   RUNG wire#w1
      R_Coil( %DB60.DBX2.7 )
   END_RUNG
   RUNG wire#w1
      R_Coil( %DB60.DBX3.0 )
   END_RUNG
   RUNG wire#w1
      R_Coil( %DB60.DBX3.1 )
   END_RUNG
   RUNG wire#w1
      R_Coil( %DB60.DBX3.2 )
   END_RUNG
   RUNG wire#w1
      R_Coil( %DB60.DBX3.3 )
   END_RUNG
   RUNG wire#w1
      R_Coil( %DB60.DBX3.4 )
   END_RUNG
   RUNG wire#w1
      R_Coil( %DB60.DBX3.5 )
   END_RUNG
   RUNG wire#w1
      R_Coil( %DB60.DBX3.6 )
   END_RUNG
   RUNG wire#w1
      R_Coil( %DB60.DBX3.7 )
   END_RUNG
   RUNG wire#w1
      R_Coil( %DB60.DBX4.0 )
   END_RUNG
   RUNG wire#w1
      R_Coil( %DB60.DBX4.1 )
   END_RUNG
   RUNG wire#w1
      R_Coil( %DB60.DBX4.2 )
   END_RUNG
   RUNG wire#w1
      R_Coil( %DB60.DBX4.3 )
   END_RUNG
   RUNG wire#w1
      R_Coil( %DB60.DBX4.4 )
   END_RUNG
   RUNG wire#w1
      R_Coil( %DB60.DBX4.5 )
   END_RUNG
   RUNG wire#w1
      R_Coil( %DB60.DBX4.6 )
   END_RUNG
   RUNG wire#w1
      R_Coil( %DB60.DBX4.7 )
   END_RUNG
   RUNG wire#w1
      R_Coil( %DB60.DBX5.0 )
   END_RUNG
   RUNG wire#w1
      R_Coil( %DB60.DBX5.1 )
   END_RUNG
   RUNG wire#w1
      R_Coil( %DB60.DBX5.2 )
   END_RUNG
   RUNG wire#w1
      R_Coil( %DB60.DBX5.3 )
   END_RUNG
   RUNG wire#w1
      R_Coil( %DB60.DBX5.4 )
   END_RUNG
   RUNG wire#w1
      R_Coil( %DB60.DBX5.5 )
   END_RUNG
   RUNG wire#w1
      R_Coil( %DB60.DBX5.6 )
   END_RUNG
   RUNG wire#w1
      R_Coil( %DB60.DBX5.7 )
   END_RUNG
   RUNG wire#w1
      R_Coil( %DB60.DBX6.0 )
   END_RUNG
   RUNG wire#w1
      R_Coil( %DB60.DBX6.1 )
   END_RUNG
   RUNG wire#w1
      R_Coil( %DB60.DBX6.2 )
   END_RUNG
   RUNG wire#w1
      R_Coil( %DB60.DBX6.3 )
   END_RUNG
   RUNG wire#w1
      R_Coil( %DB60.DBX6.4 )
   END_RUNG
   RUNG wire#w1
      R_Coil( %DB60.DBX6.5 )
   END_RUNG
   RUNG wire#w1
      R_Coil( %DB60.DBX6.6 )
   END_RUNG
   RUNG wire#w1
      R_Coil( %DB60.DBX6.7 )
   END_RUNG
   RUNG wire#w1
      R_Coil( %DB60.DBX7.0 )
   END_RUNG
   RUNG wire#w1
      R_Coil( %DB60.DBX7.1 )
   END_RUNG
   RUNG wire#w1
      R_Coil( %DB60.DBX7.2 )
   END_RUNG
   RUNG wire#w1
      R_Coil( %DB60.DBX7.3 )
   END_RUNG
   RUNG wire#w1
      R_Coil( %DB60.DBX7.4 )
   END_RUNG
   RUNG wire#w1
      R_Coil( %DB60.DBX7.5 )
   END_RUNG
   RUNG wire#w1
      R_Coil( %DB60.DBX7.6 )
   END_RUNG
   RUNG wire#w1
      R_Coil( %DB60.DBX7.7 )
   END_RUNG
   // the same network as SCL:
   IF "50_CMND_DATA".Alarm_Reset THEN
       %DB60.DBX0.0 := FALSE;
       %DB60.DBX0.1 := FALSE;
       %DB60.DBX0.2 := FALSE;
       %DB60.DBX0.3 := FALSE;
       %DB60.DBX0.4 := FALSE;
       %DB60.DBX0.5 := FALSE;
       %DB60.DBX0.6 := FALSE;
       %DB60.DBX0.7 := FALSE;
       %DB60.DBX1.0 := FALSE;
       %DB60.DBX1.1 := FALSE;
       %DB60.DBX1.2 := FALSE;
       %DB60.DBX1.3 := FALSE;
       %DB60.DBX1.4 := FALSE;
       %DB60.DBX1.5 := FALSE;
       %DB60.DBX1.6 := FALSE;
       %DB60.DBX1.7 := FALSE;
       %DB60.DBX2.0 := FALSE;
       %DB60.DBX2.1 := FALSE;
       %DB60.DBX2.2 := FALSE;
       %DB60.DBX2.3 := FALSE;
       %DB60.DBX2.4 := FALSE;
       %DB60.DBX2.5 := FALSE;
       %DB60.DBX2.6 := FALSE;
       %DB60.DBX2.7 := FALSE;
       %DB60.DBX3.0 := FALSE;
       %DB60.DBX3.1 := FALSE;
       %DB60.DBX3.2 := FALSE;
       %DB60.DBX3.3 := FALSE;
       %DB60.DBX3.4 := FALSE;
       %DB60.DBX3.5 := FALSE;
       %DB60.DBX3.6 := FALSE;
       %DB60.DBX3.7 := FALSE;
       %DB60.DBX4.0 := FALSE;
       %DB60.DBX4.1 := FALSE;
       %DB60.DBX4.2 := FALSE;
       %DB60.DBX4.3 := FALSE;
       %DB60.DBX4.4 := FALSE;
       %DB60.DBX4.5 := FALSE;
       %DB60.DBX4.6 := FALSE;
       %DB60.DBX4.7 := FALSE;
       %DB60.DBX5.0 := FALSE;
       %DB60.DBX5.1 := FALSE;
       %DB60.DBX5.2 := FALSE;
       %DB60.DBX5.3 := FALSE;
       %DB60.DBX5.4 := FALSE;
       %DB60.DBX5.5 := FALSE;
       %DB60.DBX5.6 := FALSE;
       %DB60.DBX5.7 := FALSE;
       %DB60.DBX6.0 := FALSE;
       %DB60.DBX6.1 := FALSE;
       %DB60.DBX6.2 := FALSE;
       %DB60.DBX6.3 := FALSE;
       %DB60.DBX6.4 := FALSE;
       %DB60.DBX6.5 := FALSE;
       %DB60.DBX6.6 := FALSE;
       %DB60.DBX6.7 := FALSE;
       %DB60.DBX7.0 := FALSE;
       %DB60.DBX7.1 := FALSE;
       %DB60.DBX7.2 := FALSE;
       %DB60.DBX7.3 := FALSE;
       %DB60.DBX7.4 := FALSE;
       %DB60.DBX7.5 := FALSE;
       %DB60.DBX7.6 := FALSE;
       %DB60.DBX7.7 := FALSE;
   END_IF;
END_REGION

REGION Network 34: Alarm Present
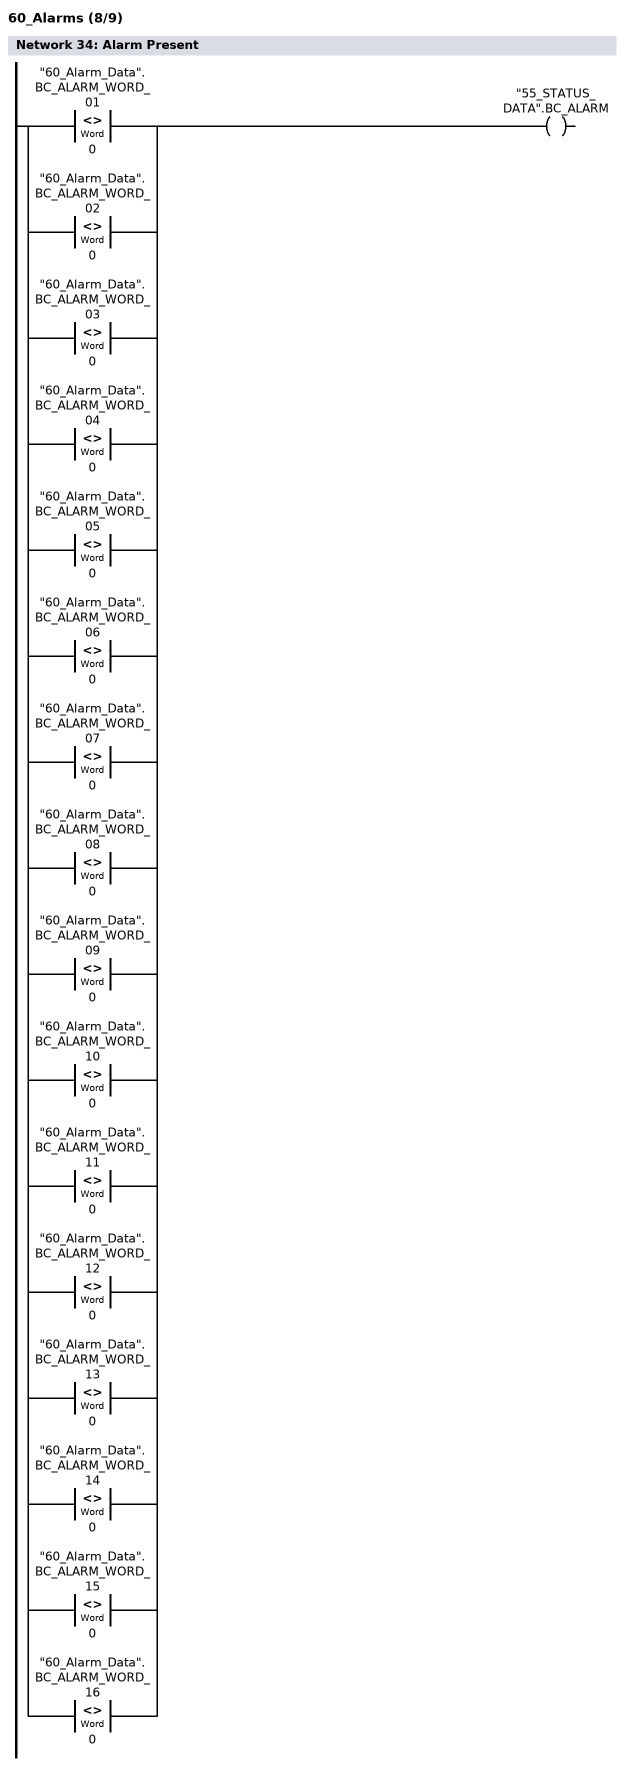
   RUNG wire#powerrail
      { S7_Templates := "SrcType := Word" } NE_Contact(in1 := "60_Alarm_Data".BC_ALARM_WORD_01, in2 := 0)
      wire#w1
      Coil( "55_STATUS_DATA".BC_ALARM )
   END_RUNG
   RUNG wire#powerrail
      { S7_Templates := "SrcType := Word" } NE_Contact(in1 := "60_Alarm_Data".BC_ALARM_WORD_02, in2 := 0)
   END_RUNG wire#w1
   RUNG wire#powerrail
      { S7_Templates := "SrcType := Word" } NE_Contact(in1 := "60_Alarm_Data".BC_ALARM_WORD_03, in2 := 0)
   END_RUNG wire#w1
   RUNG wire#powerrail
      { S7_Templates := "SrcType := Word" } NE_Contact(in1 := "60_Alarm_Data".BC_ALARM_WORD_04, in2 := 0)
   END_RUNG wire#w1
   RUNG wire#powerrail
      { S7_Templates := "SrcType := Word" } NE_Contact(in1 := "60_Alarm_Data".BC_ALARM_WORD_05, in2 := 0)
   END_RUNG wire#w1
   RUNG wire#powerrail
      { S7_Templates := "SrcType := Word" } NE_Contact(in1 := "60_Alarm_Data".BC_ALARM_WORD_06, in2 := 0)
   END_RUNG wire#w1
   RUNG wire#powerrail
      { S7_Templates := "SrcType := Word" } NE_Contact(in1 := "60_Alarm_Data".BC_ALARM_WORD_07, in2 := 0)
   END_RUNG wire#w1
   RUNG wire#powerrail
      { S7_Templates := "SrcType := Word" } NE_Contact(in1 := "60_Alarm_Data".BC_ALARM_WORD_08, in2 := 0)
   END_RUNG wire#w1
   RUNG wire#powerrail
      { S7_Templates := "SrcType := Word" } NE_Contact(in1 := "60_Alarm_Data".BC_ALARM_WORD_09, in2 := 0)
   END_RUNG wire#w1
   RUNG wire#powerrail
      { S7_Templates := "SrcType := Word" } NE_Contact(in1 := "60_Alarm_Data".BC_ALARM_WORD_10, in2 := 0)
   END_RUNG wire#w1
   RUNG wire#powerrail
      { S7_Templates := "SrcType := Word" } NE_Contact(in1 := "60_Alarm_Data".BC_ALARM_WORD_11, in2 := 0)
   END_RUNG wire#w1
   RUNG wire#powerrail
      { S7_Templates := "SrcType := Word" } NE_Contact(in1 := "60_Alarm_Data".BC_ALARM_WORD_12, in2 := 0)
   END_RUNG wire#w1
   RUNG wire#powerrail
      { S7_Templates := "SrcType := Word" } NE_Contact(in1 := "60_Alarm_Data".BC_ALARM_WORD_13, in2 := 0)
   END_RUNG wire#w1
   RUNG wire#powerrail
      { S7_Templates := "SrcType := Word" } NE_Contact(in1 := "60_Alarm_Data".BC_ALARM_WORD_14, in2 := 0)
   END_RUNG wire#w1
   RUNG wire#powerrail
      { S7_Templates := "SrcType := Word" } NE_Contact(in1 := "60_Alarm_Data".BC_ALARM_WORD_15, in2 := 0)
   END_RUNG wire#w1
   RUNG wire#powerrail
      { S7_Templates := "SrcType := Word" } NE_Contact(in1 := "60_Alarm_Data".BC_ALARM_WORD_16, in2 := 0)
   END_RUNG wire#w1
   // the same network as SCL:
   "55_STATUS_DATA".BC_ALARM := ("60_Alarm_Data".BC_ALARM_WORD_01 <> 0) OR ("60_Alarm_Data".BC_ALARM_WORD_02 <> 0) OR ("60_Alarm_Data".BC_ALARM_WORD_03 <> 0) OR ("60_Alarm_Data".BC_ALARM_WORD_04 <> 0) OR ("60_Alarm_Data".BC_ALARM_WORD_05 <> 0) OR ("60_Alarm_Data".BC_ALARM_WORD_06 <> 0) OR ("60_Alarm_Data".BC_ALARM_WORD_07 <> 0) OR ("60_Alarm_Data".BC_ALARM_WORD_08 <> 0) OR ("60_Alarm_Data".BC_ALARM_WORD_09 <> 0) OR ("60_Alarm_Data".BC_ALARM_WORD_10 <> 0) OR ("60_Alarm_Data".BC_ALARM_WORD_11 <> 0) OR ("60_Alarm_Data".BC_ALARM_WORD_12 <> 0) OR ("60_Alarm_Data".BC_ALARM_WORD_13 <> 0) OR ("60_Alarm_Data".BC_ALARM_WORD_14 <> 0) OR ("60_Alarm_Data".BC_ALARM_WORD_15 <> 0) OR ("60_Alarm_Data".BC_ALARM_WORD_16 <> 0);
END_REGION

REGION Network 35: Alarm present
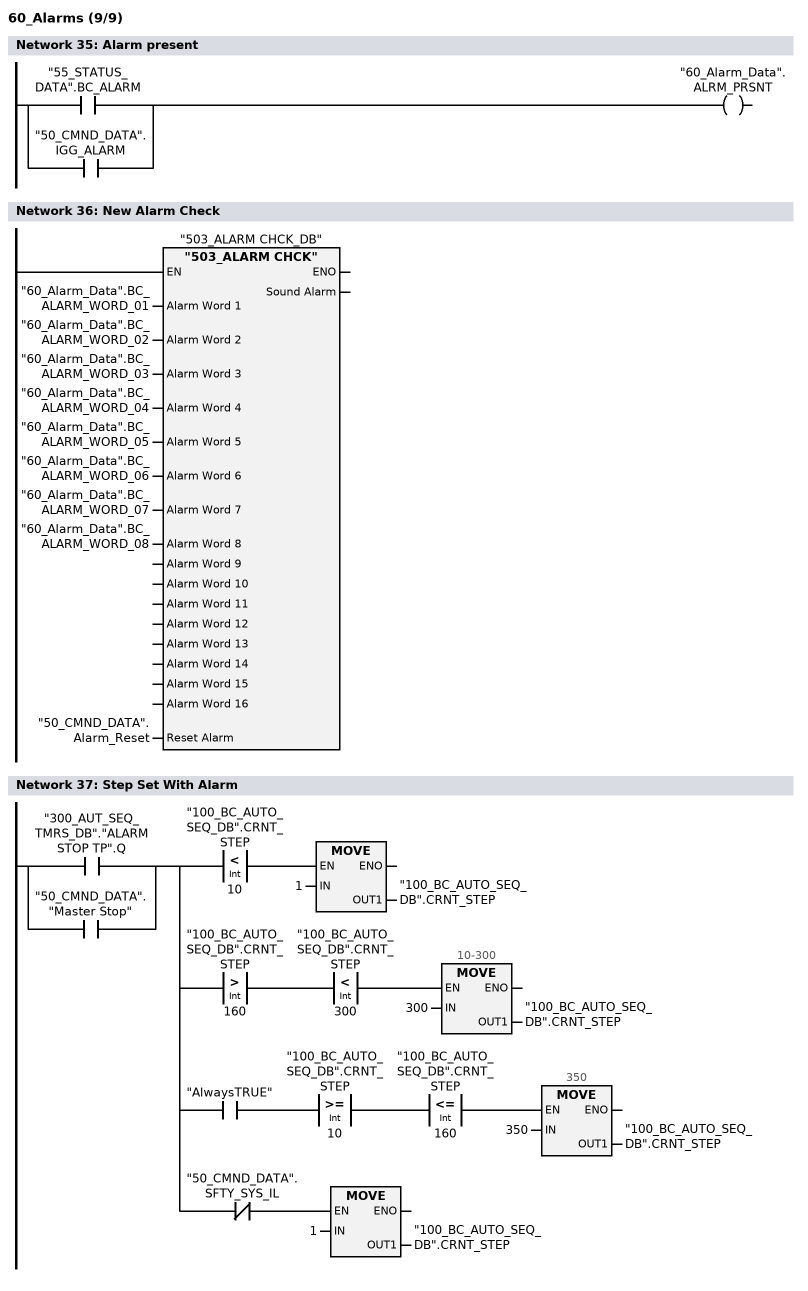
   RUNG wire#powerrail
      Contact( "55_STATUS_DATA".BC_ALARM )
      wire#w1
      Coil( "60_Alarm_Data".ALRM_PRSNT )
   END_RUNG
   RUNG wire#powerrail
      Contact( "50_CMND_DATA".IGG_ALARM )
   END_RUNG wire#w1
   // the same network as SCL:
   "60_Alarm_Data".ALRM_PRSNT := "55_STATUS_DATA".BC_ALARM OR "50_CMND_DATA".IGG_ALARM;
END_REGION

REGION Network 36: New Alarm Check
   RUNG wire#powerrail
      "503_ALARM CHCK_DB"("Alarm Word 1" := "60_Alarm_Data".BC_ALARM_WORD_01, "Alarm Word 2" := "60_Alarm_Data".BC_ALARM_WORD_02, "Alarm Word 3" := "60_Alarm_Data".BC_ALARM_WORD_03, "Alarm Word 4" := "60_Alarm_Data".BC_ALARM_WORD_04, "Alarm Word 5" := "60_Alarm_Data".BC_ALARM_WORD_05, "Alarm Word 6" := "60_Alarm_Data".BC_ALARM_WORD_06, "Alarm Word 7" := "60_Alarm_Data".BC_ALARM_WORD_07, "Alarm Word 8" := "60_Alarm_Data".BC_ALARM_WORD_08, "Alarm Word 9" :=, "Alarm Word 10" :=, "Alarm Word 11" :=, "Alarm Word 12" :=, "Alarm Word 13" :=, "Alarm Word 14" :=, "Alarm Word 15" :=, "Alarm Word 16" :=, "Reset Alarm" := "50_CMND_DATA".Alarm_Reset, "Sound Alarm" =>)
   END_RUNG
   // the same network as SCL:
   "503_ALARM CHCK_DB"("Alarm Word 1" := "60_Alarm_Data".BC_ALARM_WORD_01,   // "503_ALARM CHCK"
                       "Alarm Word 2" := "60_Alarm_Data".BC_ALARM_WORD_02,
                       "Alarm Word 3" := "60_Alarm_Data".BC_ALARM_WORD_03,
                       "Alarm Word 4" := "60_Alarm_Data".BC_ALARM_WORD_04,
                       "Alarm Word 5" := "60_Alarm_Data".BC_ALARM_WORD_05,
                       "Alarm Word 6" := "60_Alarm_Data".BC_ALARM_WORD_06,
                       "Alarm Word 7" := "60_Alarm_Data".BC_ALARM_WORD_07,
                       "Alarm Word 8" := "60_Alarm_Data".BC_ALARM_WORD_08,
                       "Reset Alarm" := "50_CMND_DATA".Alarm_Reset);
END_REGION

REGION Network 37: Step Set With Alarm
   RUNG wire#powerrail
      Contact( "300_AUT_SEQ_TMRS_DB"."ALARM STOP TP".Q )
      wire#w1
      { S7_Templates := "SrcType := Int" } LT_Contact(in1 := "100_BC_AUTO_SEQ_DB".CRNT_STEP, in2 := 10)
      Move(in := 1, out1 => "100_BC_AUTO_SEQ_DB".CRNT_STEP)
   END_RUNG
   RUNG wire#powerrail
      Contact( "50_CMND_DATA"."Master Stop" )
   END_RUNG wire#w1
   RUNG wire#w1
      { S7_Templates := "SrcType := Int" } GT_Contact(in1 := "100_BC_AUTO_SEQ_DB".CRNT_STEP, in2 := 160)
      { S7_Templates := "SrcType := Int" } LT_Contact(in1 := "100_BC_AUTO_SEQ_DB".CRNT_STEP, in2 := 300)
      Move(in := 300, out1 => "100_BC_AUTO_SEQ_DB".CRNT_STEP)   // 10-300
   END_RUNG
   RUNG wire#w1
      Contact( "AlwaysTRUE" )
      { S7_Templates := "SrcType := Int" } GE_Contact(in1 := "100_BC_AUTO_SEQ_DB".CRNT_STEP, in2 := 10)
      { S7_Templates := "SrcType := Int" } LE_Contact(in1 := "100_BC_AUTO_SEQ_DB".CRNT_STEP, in2 := 160)
      Move(in := 350, out1 => "100_BC_AUTO_SEQ_DB".CRNT_STEP)   // 350
   END_RUNG
   RUNG wire#w1
      I_Contact( "50_CMND_DATA".SFTY_SYS_IL )
      Move(in := 1, out1 => "100_BC_AUTO_SEQ_DB".CRNT_STEP)
   END_RUNG
   // the same network as SCL:
   #_w1 := "300_AUT_SEQ_TMRS_DB"."ALARM STOP TP".Q OR "50_CMND_DATA"."Master Stop";
   IF #_w1 AND ("100_BC_AUTO_SEQ_DB".CRNT_STEP < 10) THEN "100_BC_AUTO_SEQ_DB".CRNT_STEP := 1; END_IF;
   IF #_w1 AND ("100_BC_AUTO_SEQ_DB".CRNT_STEP > 160) AND ("100_BC_AUTO_SEQ_DB".CRNT_STEP < 300) THEN
       "100_BC_AUTO_SEQ_DB".CRNT_STEP := 300;   // 10-300
   END_IF;
   IF #_w1 AND "AlwaysTRUE" AND ("100_BC_AUTO_SEQ_DB".CRNT_STEP >= 10) AND ("100_BC_AUTO_SEQ_DB".CRNT_STEP <= 160) THEN
       "100_BC_AUTO_SEQ_DB".CRNT_STEP := 350;   // 350
   END_IF;
   IF #_w1 AND NOT "50_CMND_DATA".SFTY_SYS_IL THEN "100_BC_AUTO_SEQ_DB".CRNT_STEP := 1; END_IF;
END_REGION
END_FUNCTION

FUNCTION "62_Warnings" : Void   // FC62, LAD
TITLE = Warning Processing
{ S7_Optimized_Access := 'TRUE' }
AUTHOR : JRS
VERSION : 0.1
// To warning conditions
   VAR_TEMP   // added for the SCL form of the ladder/FBD networks
      _w1 : Bool;
   END_VAR
BEGIN

REGION Network 1: DB62 WORD_1 =PIT204 Fuel Oil pessure transmitter
   // BC_WARNING_WORD_01 BIT 1/2/3/4
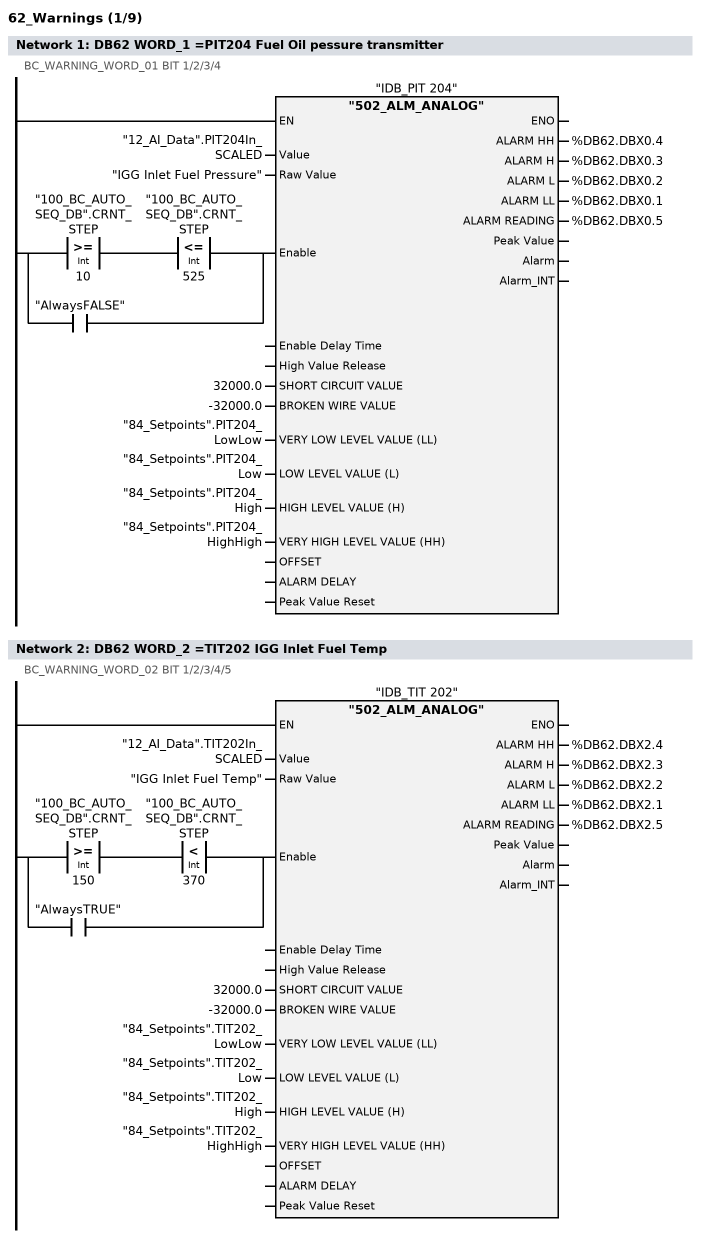
   RUNG wire#powerrail
      "IDB_PIT 204"(Enable := wire#w1, Value := "12_AI_Data".PIT204In_SCALED, "Raw Value" := "IGG Inlet Fuel Pressure", "SHORT CIRCUIT VALUE" := 32000.0, "BROKEN WIRE VALUE" := -32000.0, "VERY LOW LEVEL VALUE (LL)" := "84_Setpoints".PIT204_LowLow, "LOW LEVEL VALUE (L)" := "84_Setpoints".PIT204_Low, "HIGH LEVEL VALUE (H)" := "84_Setpoints".PIT204_High, "VERY HIGH LEVEL VALUE (HH)" := "84_Setpoints".PIT204_HighHigh, OFFSET :=, "ALARM DELAY" :=, "Peak Value Reset" :=, "ALARM HH" => %DB62.DBX0.4, "ALARM H" => %DB62.DBX0.3, "ALARM L" => %DB62.DBX0.2, "ALARM LL" => %DB62.DBX0.1, "ALARM READING" => %DB62.DBX0.5, "Peak Value" =>, Alarm =>, Alarm_INT =>, "Enable Delay Time" :=, "High Value Release" :=)
   END_RUNG
   RUNG wire#powerrail
      { S7_Templates := "SrcType := Int" } GE_Contact(in1 := "100_BC_AUTO_SEQ_DB".CRNT_STEP, in2 := 10)
      { S7_Templates := "SrcType := Int" } LE_Contact(in1 := "100_BC_AUTO_SEQ_DB".CRNT_STEP, in2 := 525)
   END_RUNG wire#w1
   RUNG wire#powerrail
      Contact( "AlwaysFALSE" )
   END_RUNG wire#w1
   // the same network as SCL:
   "IDB_PIT 204"(Value := "12_AI_Data".PIT204In_SCALED,   // "502_ALM_ANALOG"
                 "Raw Value" := "IGG Inlet Fuel Pressure",
                 Enable := (("100_BC_AUTO_SEQ_DB".CRNT_STEP >= 10) AND ("100_BC_AUTO_SEQ_DB".CRNT_STEP <= 525)) OR "AlwaysFALSE",
                 "SHORT CIRCUIT VALUE" := 32000.0,
                 "BROKEN WIRE VALUE" := -32000.0,
                 "VERY LOW LEVEL VALUE (LL)" := "84_Setpoints".PIT204_LowLow,
                 "LOW LEVEL VALUE (L)" := "84_Setpoints".PIT204_Low,
                 "HIGH LEVEL VALUE (H)" := "84_Setpoints".PIT204_High,
                 "VERY HIGH LEVEL VALUE (HH)" := "84_Setpoints".PIT204_HighHigh,
                 "ALARM HH" => %DB62.DBX0.4,
                 "ALARM H" => %DB62.DBX0.3,
                 "ALARM L" => %DB62.DBX0.2,
                 "ALARM LL" => %DB62.DBX0.1,
                 "ALARM READING" => %DB62.DBX0.5);
END_REGION

REGION Network 2: DB62 WORD_2 =TIT202 IGG Inlet Fuel Temp
   // BC_WARNING_WORD_02 BIT 1/2/3/4/5
   RUNG wire#powerrail
      "IDB_TIT 202"(Enable := wire#w1, Value := "12_AI_Data".TIT202In_SCALED, "Raw Value" := "IGG Inlet Fuel Temp", "SHORT CIRCUIT VALUE" := 32000.0, "BROKEN WIRE VALUE" := -32000.0, "VERY LOW LEVEL VALUE (LL)" := "84_Setpoints".TIT202_LowLow, "LOW LEVEL VALUE (L)" := "84_Setpoints".TIT202_Low, "HIGH LEVEL VALUE (H)" := "84_Setpoints".TIT202_High, "VERY HIGH LEVEL VALUE (HH)" := "84_Setpoints".TIT202_HighHigh, OFFSET :=, "ALARM DELAY" :=, "Peak Value Reset" :=, "ALARM HH" => %DB62.DBX2.4, "ALARM H" => %DB62.DBX2.3, "ALARM L" => %DB62.DBX2.2, "ALARM LL" => %DB62.DBX2.1, "ALARM READING" => %DB62.DBX2.5, "Peak Value" =>, Alarm =>, Alarm_INT =>, "Enable Delay Time" :=, "High Value Release" :=)
   END_RUNG
   RUNG wire#powerrail
      { S7_Templates := "SrcType := Int" } GE_Contact(in1 := "100_BC_AUTO_SEQ_DB".CRNT_STEP, in2 := 150)
      { S7_Templates := "SrcType := Int" } LT_Contact(in1 := "100_BC_AUTO_SEQ_DB".CRNT_STEP, in2 := 370)
   END_RUNG wire#w1
   RUNG wire#powerrail
      Contact( "AlwaysTRUE" )
   END_RUNG wire#w1
   // the same network as SCL:
   "IDB_TIT 202"(Value := "12_AI_Data".TIT202In_SCALED,   // "502_ALM_ANALOG"
                 "Raw Value" := "IGG Inlet Fuel Temp",
                 Enable := (("100_BC_AUTO_SEQ_DB".CRNT_STEP >= 150) AND ("100_BC_AUTO_SEQ_DB".CRNT_STEP < 370)) OR "AlwaysTRUE",
                 "SHORT CIRCUIT VALUE" := 32000.0,
                 "BROKEN WIRE VALUE" := -32000.0,
                 "VERY LOW LEVEL VALUE (LL)" := "84_Setpoints".TIT202_LowLow,
                 "LOW LEVEL VALUE (L)" := "84_Setpoints".TIT202_Low,
                 "HIGH LEVEL VALUE (H)" := "84_Setpoints".TIT202_High,
                 "VERY HIGH LEVEL VALUE (HH)" := "84_Setpoints".TIT202_HighHigh,
                 "ALARM HH" => %DB62.DBX2.4,
                 "ALARM H" => %DB62.DBX2.3,
                 "ALARM L" => %DB62.DBX2.2,
                 "ALARM LL" => %DB62.DBX2.1,
                 "ALARM READING" => %DB62.DBX2.5);
END_REGION

REGION Network 3: DB62 WORD_3 =PIT205 IGG Main Fuel Pressure
   // BC_WARNING_WORD_03
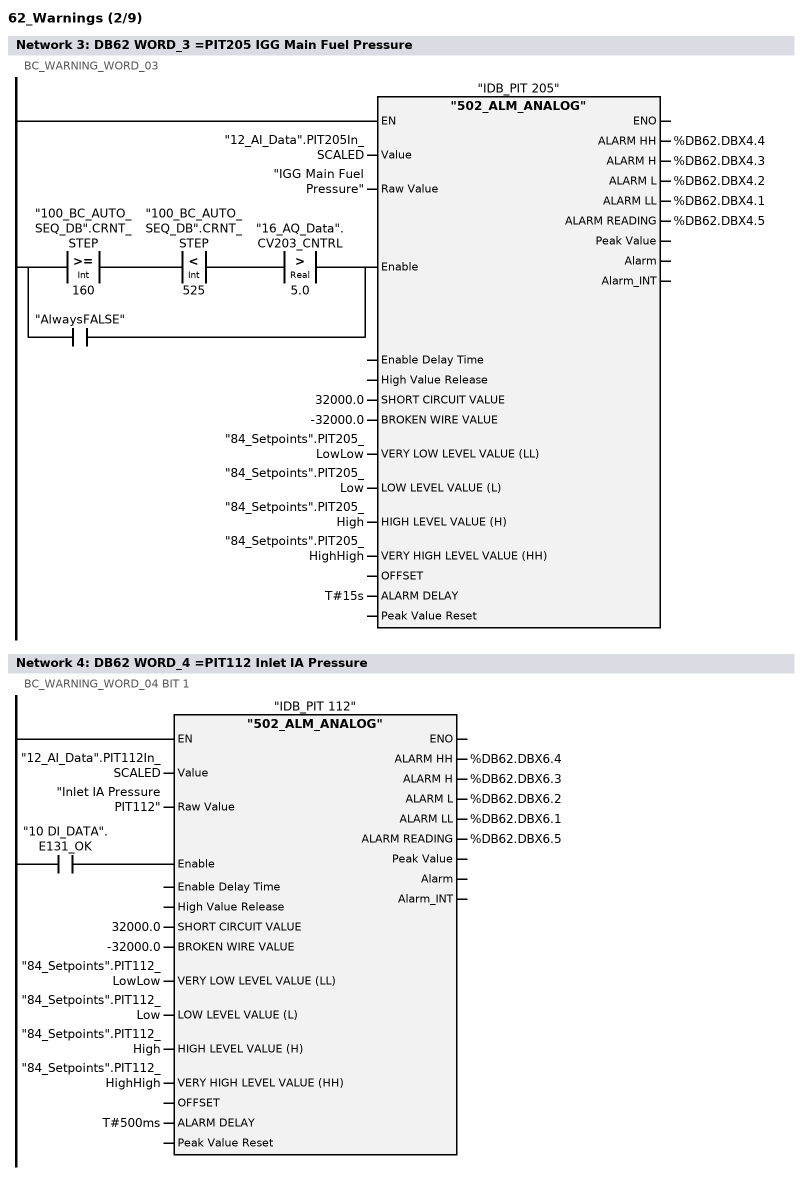
   RUNG wire#powerrail
      "IDB_PIT 205"(Enable := wire#w1, Value := "12_AI_Data".PIT205In_SCALED, "Raw Value" := "IGG Main Fuel Pressure", "SHORT CIRCUIT VALUE" := 32000.0, "BROKEN WIRE VALUE" := -32000.0, "VERY LOW LEVEL VALUE (LL)" := "84_Setpoints".PIT205_LowLow, "LOW LEVEL VALUE (L)" := "84_Setpoints".PIT205_Low, "HIGH LEVEL VALUE (H)" := "84_Setpoints".PIT205_High, "VERY HIGH LEVEL VALUE (HH)" := "84_Setpoints".PIT205_HighHigh, OFFSET :=, "ALARM DELAY" := T#15s, "Peak Value Reset" :=, "ALARM HH" => %DB62.DBX4.4, "ALARM H" => %DB62.DBX4.3, "ALARM L" => %DB62.DBX4.2, "ALARM LL" => %DB62.DBX4.1, "ALARM READING" => %DB62.DBX4.5, "Peak Value" =>, Alarm =>, Alarm_INT =>, "Enable Delay Time" :=, "High Value Release" :=)
   END_RUNG
   RUNG wire#powerrail
      { S7_Templates := "SrcType := Int" } GE_Contact(in1 := "100_BC_AUTO_SEQ_DB".CRNT_STEP, in2 := 160)
      { S7_Templates := "SrcType := Int" } LT_Contact(in1 := "100_BC_AUTO_SEQ_DB".CRNT_STEP, in2 := 525)
      { S7_Templates := "SrcType := Real" } GT_Contact(in1 := "16_AQ_Data".CV203_CNTRL, in2 := 5.0)
   END_RUNG wire#w1
   RUNG wire#powerrail
      Contact( "AlwaysFALSE" )
   END_RUNG wire#w1
   // the same network as SCL:
   "IDB_PIT 205"(Value := "12_AI_Data".PIT205In_SCALED,   // "502_ALM_ANALOG"
                 "Raw Value" := "IGG Main Fuel Pressure",
                 Enable := (("100_BC_AUTO_SEQ_DB".CRNT_STEP >= 160) AND ("100_BC_AUTO_SEQ_DB".CRNT_STEP < 525) AND ("16_AQ_Data".CV203_CNTRL > 5.0)) OR "AlwaysFALSE",
                 "SHORT CIRCUIT VALUE" := 32000.0,
                 "BROKEN WIRE VALUE" := -32000.0,
                 "VERY LOW LEVEL VALUE (LL)" := "84_Setpoints".PIT205_LowLow,
                 "LOW LEVEL VALUE (L)" := "84_Setpoints".PIT205_Low,
                 "HIGH LEVEL VALUE (H)" := "84_Setpoints".PIT205_High,
                 "VERY HIGH LEVEL VALUE (HH)" := "84_Setpoints".PIT205_HighHigh,
                 "ALARM DELAY" := T#15s,
                 "ALARM HH" => %DB62.DBX4.4,
                 "ALARM H" => %DB62.DBX4.3,
                 "ALARM L" => %DB62.DBX4.2,
                 "ALARM LL" => %DB62.DBX4.1,
                 "ALARM READING" => %DB62.DBX4.5);
END_REGION

REGION Network 4: DB62 WORD_4 =PIT112 Inlet IA Pressure
   // BC_WARNING_WORD_04 BIT 1
   RUNG wire#powerrail
      "IDB_PIT 112"(Enable := wire#w1, Value := "12_AI_Data".PIT112In_SCALED, "Raw Value" := "Inlet IA Pressure PIT112", "SHORT CIRCUIT VALUE" := 32000.0, "BROKEN WIRE VALUE" := -32000.0, "VERY LOW LEVEL VALUE (LL)" := "84_Setpoints".PIT112_LowLow, "LOW LEVEL VALUE (L)" := "84_Setpoints".PIT112_Low, "HIGH LEVEL VALUE (H)" := "84_Setpoints".PIT112_High, "VERY HIGH LEVEL VALUE (HH)" := "84_Setpoints".PIT112_HighHigh, OFFSET :=, "ALARM DELAY" := T#500ms, "Peak Value Reset" :=, "ALARM HH" => %DB62.DBX6.4, "ALARM H" => %DB62.DBX6.3, "ALARM L" => %DB62.DBX6.2, "ALARM LL" => %DB62.DBX6.1, "ALARM READING" => %DB62.DBX6.5, "Peak Value" =>, Alarm =>, Alarm_INT =>, "Enable Delay Time" :=, "High Value Release" :=)
   END_RUNG
   RUNG wire#powerrail
      Contact( "10 DI_DATA".E131_OK )
   END_RUNG wire#w1
   // the same network as SCL:
   "IDB_PIT 112"(Value := "12_AI_Data".PIT112In_SCALED,   // "502_ALM_ANALOG"
                 "Raw Value" := "Inlet IA Pressure PIT112",
                 Enable := "10 DI_DATA".E131_OK,
                 "SHORT CIRCUIT VALUE" := 32000.0,
                 "BROKEN WIRE VALUE" := -32000.0,
                 "VERY LOW LEVEL VALUE (LL)" := "84_Setpoints".PIT112_LowLow,
                 "LOW LEVEL VALUE (L)" := "84_Setpoints".PIT112_Low,
                 "HIGH LEVEL VALUE (H)" := "84_Setpoints".PIT112_High,
                 "VERY HIGH LEVEL VALUE (HH)" := "84_Setpoints".PIT112_HighHigh,
                 "ALARM DELAY" := T#500ms,
                 "ALARM HH" => %DB62.DBX6.4,
                 "ALARM H" => %DB62.DBX6.3,
                 "ALARM L" => %DB62.DBX6.2,
                 "ALARM LL" => %DB62.DBX6.1,
                 "ALARM READING" => %DB62.DBX6.5);
END_REGION

REGION Network 5: DB62 WORD_5 =PIT113 IGG Main Atom Air Pressure
   // BC_WARNING_WORD_05
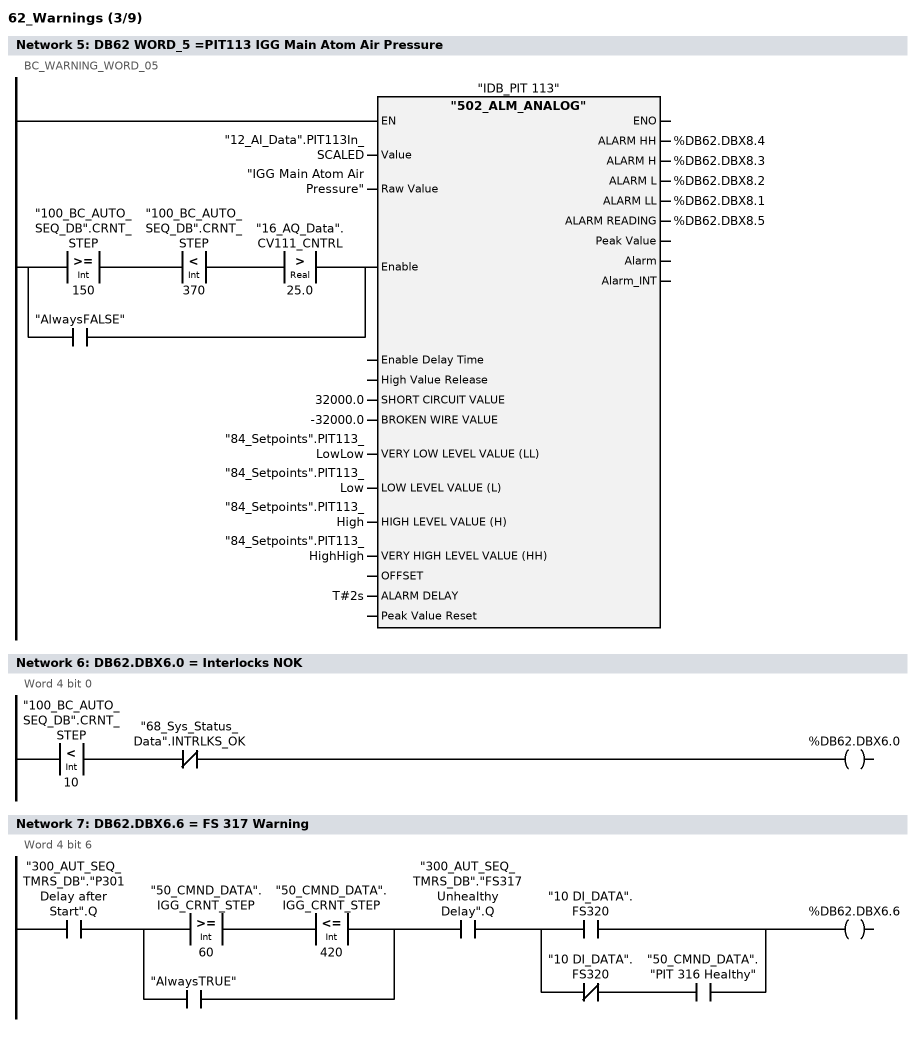
   RUNG wire#powerrail
      "IDB_PIT 113"(Enable := wire#w1, Value := "12_AI_Data".PIT113In_SCALED, "Raw Value" := "IGG Main Atom Air Pressure", "SHORT CIRCUIT VALUE" := 32000.0, "BROKEN WIRE VALUE" := -32000.0, "VERY LOW LEVEL VALUE (LL)" := "84_Setpoints".PIT113_LowLow, "LOW LEVEL VALUE (L)" := "84_Setpoints".PIT113_Low, "HIGH LEVEL VALUE (H)" := "84_Setpoints".PIT113_High, "VERY HIGH LEVEL VALUE (HH)" := "84_Setpoints".PIT113_HighHigh, OFFSET :=, "ALARM DELAY" := T#2s, "Peak Value Reset" :=, "ALARM HH" => %DB62.DBX8.4, "ALARM H" => %DB62.DBX8.3, "ALARM L" => %DB62.DBX8.2, "ALARM LL" => %DB62.DBX8.1, "ALARM READING" => %DB62.DBX8.5, "Peak Value" =>, Alarm =>, Alarm_INT =>, "Enable Delay Time" :=, "High Value Release" :=)
   END_RUNG
   RUNG wire#powerrail
      { S7_Templates := "SrcType := Int" } GE_Contact(in1 := "100_BC_AUTO_SEQ_DB".CRNT_STEP, in2 := 150)
      { S7_Templates := "SrcType := Int" } LT_Contact(in1 := "100_BC_AUTO_SEQ_DB".CRNT_STEP, in2 := 370)
      { S7_Templates := "SrcType := Real" } GT_Contact(in1 := "16_AQ_Data".CV111_CNTRL, in2 := 25.0)
   END_RUNG wire#w1
   RUNG wire#powerrail
      Contact( "AlwaysFALSE" )
   END_RUNG wire#w1
   // the same network as SCL:
   "IDB_PIT 113"(Value := "12_AI_Data".PIT113In_SCALED,   // "502_ALM_ANALOG"
                 "Raw Value" := "IGG Main Atom Air Pressure",
                 Enable := (("100_BC_AUTO_SEQ_DB".CRNT_STEP >= 150) AND ("100_BC_AUTO_SEQ_DB".CRNT_STEP < 370) AND ("16_AQ_Data".CV111_CNTRL > 25.0)) OR "AlwaysFALSE",
                 "SHORT CIRCUIT VALUE" := 32000.0,
                 "BROKEN WIRE VALUE" := -32000.0,
                 "VERY LOW LEVEL VALUE (LL)" := "84_Setpoints".PIT113_LowLow,
                 "LOW LEVEL VALUE (L)" := "84_Setpoints".PIT113_Low,
                 "HIGH LEVEL VALUE (H)" := "84_Setpoints".PIT113_High,
                 "VERY HIGH LEVEL VALUE (HH)" := "84_Setpoints".PIT113_HighHigh,
                 "ALARM DELAY" := T#2s,
                 "ALARM HH" => %DB62.DBX8.4,
                 "ALARM H" => %DB62.DBX8.3,
                 "ALARM L" => %DB62.DBX8.2,
                 "ALARM LL" => %DB62.DBX8.1,
                 "ALARM READING" => %DB62.DBX8.5);
END_REGION

REGION Network 6: DB62.DBX6.0 = Interlocks NOK
   // Word 4 bit 0
   RUNG wire#powerrail
      { S7_Templates := "SrcType := Int" } LT_Contact(in1 := "100_BC_AUTO_SEQ_DB".CRNT_STEP, in2 := 10)
      I_Contact( "68_Sys_Status_Data".INTRLKS_OK )
      Coil( %DB62.DBX6.0 )
   END_RUNG
   // the same network as SCL:
   %DB62.DBX6.0 := ("100_BC_AUTO_SEQ_DB".CRNT_STEP < 10) AND NOT "68_Sys_Status_Data".INTRLKS_OK;
END_REGION

REGION Network 7: DB62.DBX6.6 = FS 317 Warning
   // Word 4 bit 6
   RUNG wire#powerrail
      Contact( "300_AUT_SEQ_TMRS_DB"."P301 Delay after Start".Q )
      wire#w1
      { S7_Templates := "SrcType := Int" } GE_Contact(in1 := "50_CMND_DATA".IGG_CRNT_STEP, in2 := 60)
      { S7_Templates := "SrcType := Int" } LE_Contact(in1 := "50_CMND_DATA".IGG_CRNT_STEP, in2 := 420)
      wire#w2
      Contact( "300_AUT_SEQ_TMRS_DB"."FS317 Unhealthy Delay".Q )
      wire#w3
      Contact( "10 DI_DATA".FS320 )
      wire#w4
      Coil( %DB62.DBX6.6 )
   END_RUNG
   RUNG wire#w1
      Contact( "AlwaysTRUE" )
   END_RUNG wire#w2
   RUNG wire#w3
      I_Contact( "10 DI_DATA".FS320 )
      Contact( "50_CMND_DATA"."PIT 316 Healthy" )
   END_RUNG wire#w4
   // the same network as SCL:
   %DB62.DBX6.6 := "300_AUT_SEQ_TMRS_DB"."P301 Delay after Start".Q AND ((("50_CMND_DATA".IGG_CRNT_STEP >= 60) AND ("50_CMND_DATA".IGG_CRNT_STEP <= 420)) OR "AlwaysTRUE") AND "300_AUT_SEQ_TMRS_DB"."FS317 Unhealthy Delay".Q AND ("10 DI_DATA".FS320 OR (NOT "10 DI_DATA".FS320 AND "50_CMND_DATA"."PIT 316 Healthy"));
END_REGION

REGION Network 8: DB62.DBX6.7 = FS 320 Warning
   // Word 4 bit 7
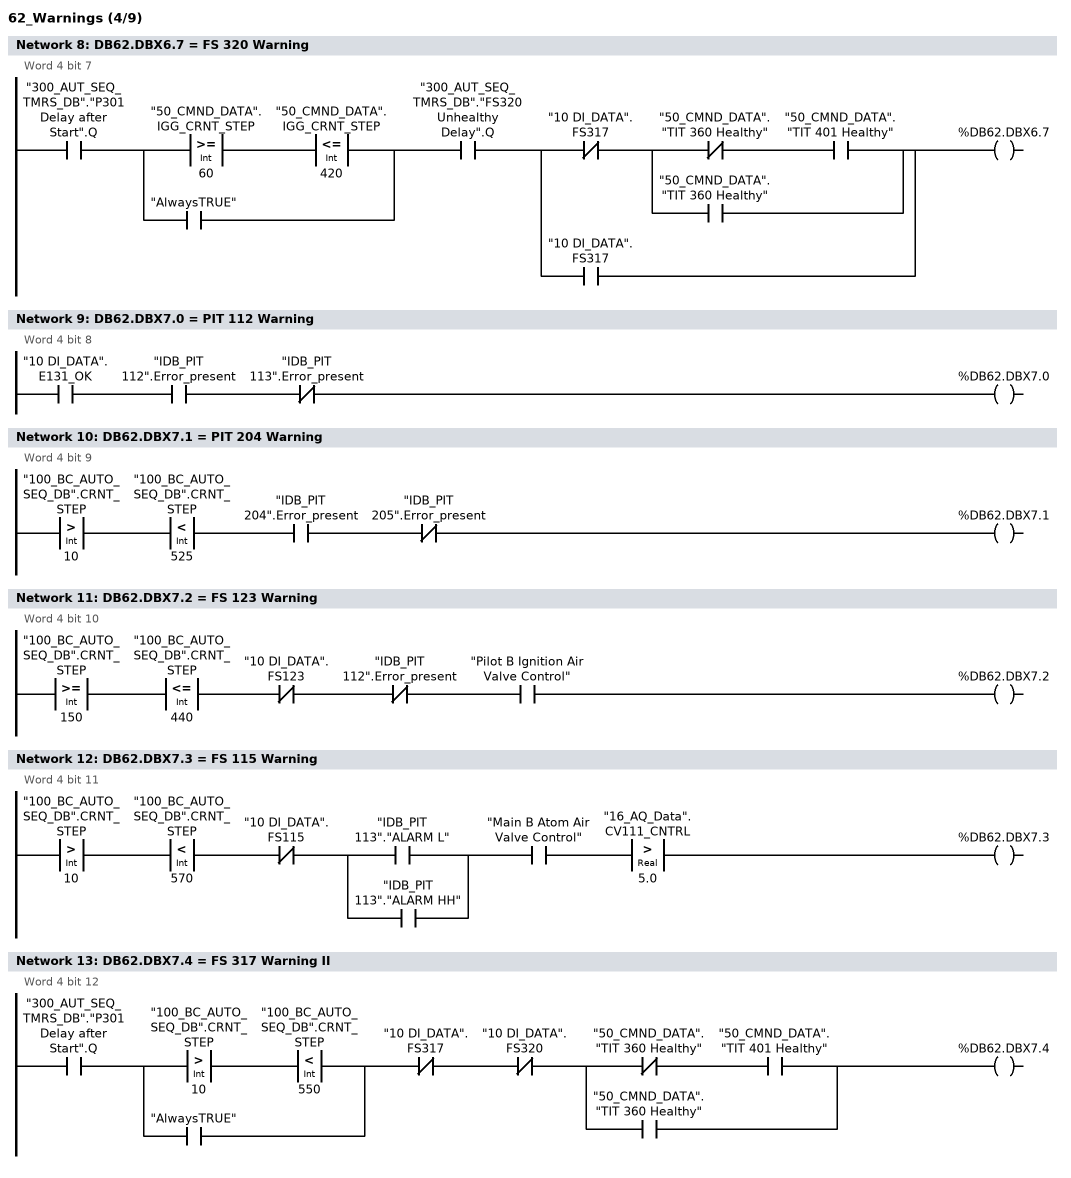
   RUNG wire#powerrail
      Contact( "300_AUT_SEQ_TMRS_DB"."P301 Delay after Start".Q )
      wire#w1
      { S7_Templates := "SrcType := Int" } GE_Contact(in1 := "50_CMND_DATA".IGG_CRNT_STEP, in2 := 60)
      { S7_Templates := "SrcType := Int" } LE_Contact(in1 := "50_CMND_DATA".IGG_CRNT_STEP, in2 := 420)
      wire#w2
      Contact( "300_AUT_SEQ_TMRS_DB"."FS320 Unhealthy Delay".Q )
      wire#w3
      I_Contact( "10 DI_DATA".FS317 )
      wire#w4
      I_Contact( "50_CMND_DATA"."TIT 360 Healthy" )
      Contact( "50_CMND_DATA"."TIT 401 Healthy" )
      wire#w5
      Coil( %DB62.DBX6.7 )
   END_RUNG
   RUNG wire#w1
      Contact( "AlwaysTRUE" )
   END_RUNG wire#w2
   RUNG wire#w4
      Contact( "50_CMND_DATA"."TIT 360 Healthy" )
   END_RUNG wire#w5
   RUNG wire#w3
      Contact( "10 DI_DATA".FS317 )
   END_RUNG wire#w5
   // the same network as SCL:
   %DB62.DBX6.7 := "300_AUT_SEQ_TMRS_DB"."P301 Delay after Start".Q AND ((("50_CMND_DATA".IGG_CRNT_STEP >= 60) AND ("50_CMND_DATA".IGG_CRNT_STEP <= 420)) OR "AlwaysTRUE") AND "300_AUT_SEQ_TMRS_DB"."FS320 Unhealthy Delay".Q AND ((NOT "10 DI_DATA".FS317 AND ((NOT "50_CMND_DATA"."TIT 360 Healthy" AND "50_CMND_DATA"."TIT 401 Healthy") OR "50_CMND_DATA"."TIT 360 Healthy")) OR "10 DI_DATA".FS317);
END_REGION

REGION Network 9: DB62.DBX7.0 = PIT 112 Warning
   // Word 4 bit 8
   RUNG wire#powerrail
      Contact( "10 DI_DATA".E131_OK )
      Contact( "IDB_PIT 112".Error_present )
      I_Contact( "IDB_PIT 113".Error_present )
      Coil( %DB62.DBX7.0 )
   END_RUNG
   // the same network as SCL:
   %DB62.DBX7.0 := "10 DI_DATA".E131_OK AND "IDB_PIT 112".Error_present AND NOT "IDB_PIT 113".Error_present;
END_REGION

REGION Network 10: DB62.DBX7.1 = PIT 204 Warning
   // Word 4 bit 9
   RUNG wire#powerrail
      { S7_Templates := "SrcType := Int" } GT_Contact(in1 := "100_BC_AUTO_SEQ_DB".CRNT_STEP, in2 := 10)
      { S7_Templates := "SrcType := Int" } LT_Contact(in1 := "100_BC_AUTO_SEQ_DB".CRNT_STEP, in2 := 525)
      Contact( "IDB_PIT 204".Error_present )
      I_Contact( "IDB_PIT 205".Error_present )
      Coil( %DB62.DBX7.1 )
   END_RUNG
   // the same network as SCL:
   %DB62.DBX7.1 := ("100_BC_AUTO_SEQ_DB".CRNT_STEP > 10) AND ("100_BC_AUTO_SEQ_DB".CRNT_STEP < 525) AND "IDB_PIT 204".Error_present AND NOT "IDB_PIT 205".Error_present;
END_REGION

REGION Network 11: DB62.DBX7.2 = FS 123 Warning
   // Word 4 bit 10
   RUNG wire#powerrail
      { S7_Templates := "SrcType := Int" } GE_Contact(in1 := "100_BC_AUTO_SEQ_DB".CRNT_STEP, in2 := 150)
      { S7_Templates := "SrcType := Int" } LE_Contact(in1 := "100_BC_AUTO_SEQ_DB".CRNT_STEP, in2 := 440)
      I_Contact( "10 DI_DATA".FS123 )
      I_Contact( "IDB_PIT 112".Error_present )
      Contact( "Pilot B Ignition Air Valve Control" )
      Coil( %DB62.DBX7.2 )
   END_RUNG
   // the same network as SCL:
   %DB62.DBX7.2 := ("100_BC_AUTO_SEQ_DB".CRNT_STEP >= 150) AND ("100_BC_AUTO_SEQ_DB".CRNT_STEP <= 440) AND NOT "10 DI_DATA".FS123 AND NOT "IDB_PIT 112".Error_present AND "Pilot B Ignition Air Valve Control";
END_REGION

REGION Network 12: DB62.DBX7.3 = FS 115 Warning
   // Word 4 bit 11
   RUNG wire#powerrail
      { S7_Templates := "SrcType := Int" } GT_Contact(in1 := "100_BC_AUTO_SEQ_DB".CRNT_STEP, in2 := 10)
      { S7_Templates := "SrcType := Int" } LT_Contact(in1 := "100_BC_AUTO_SEQ_DB".CRNT_STEP, in2 := 570)
      I_Contact( "10 DI_DATA".FS115 )
      wire#w1
      Contact( "IDB_PIT 113"."ALARM L" )
      wire#w2
      Contact( "Main B Atom Air Valve Control" )
      { S7_Templates := "SrcType := Real" } GT_Contact(in1 := "16_AQ_Data".CV111_CNTRL, in2 := 5.0)
      Coil( %DB62.DBX7.3 )
   END_RUNG
   RUNG wire#w1
      Contact( "IDB_PIT 113"."ALARM HH" )
   END_RUNG wire#w2
   // the same network as SCL:
   %DB62.DBX7.3 := ("100_BC_AUTO_SEQ_DB".CRNT_STEP > 10) AND ("100_BC_AUTO_SEQ_DB".CRNT_STEP < 570) AND NOT "10 DI_DATA".FS115 AND ("IDB_PIT 113"."ALARM L" OR "IDB_PIT 113"."ALARM HH") AND "Main B Atom Air Valve Control" AND ("16_AQ_Data".CV111_CNTRL > 5.0);
END_REGION

REGION Network 13: DB62.DBX7.4 = FS 317 Warning II
   // Word 4 bit 12
   RUNG wire#powerrail
      Contact( "300_AUT_SEQ_TMRS_DB"."P301 Delay after Start".Q )
      wire#w1
      { S7_Templates := "SrcType := Int" } GT_Contact(in1 := "100_BC_AUTO_SEQ_DB".CRNT_STEP, in2 := 10)
      { S7_Templates := "SrcType := Int" } LT_Contact(in1 := "100_BC_AUTO_SEQ_DB".CRNT_STEP, in2 := 550)
      wire#w2
      I_Contact( "10 DI_DATA".FS317 )
      I_Contact( "10 DI_DATA".FS320 )
      wire#w3
      I_Contact( "50_CMND_DATA"."TIT 360 Healthy" )
      Contact( "50_CMND_DATA"."TIT 401 Healthy" )
      wire#w4
      Coil( %DB62.DBX7.4 )
   END_RUNG
   RUNG wire#w1
      Contact( "AlwaysTRUE" )
   END_RUNG wire#w2
   RUNG wire#w3
      Contact( "50_CMND_DATA"."TIT 360 Healthy" )
   END_RUNG wire#w4
   // the same network as SCL:
   %DB62.DBX7.4 := "300_AUT_SEQ_TMRS_DB"."P301 Delay after Start".Q AND ((("100_BC_AUTO_SEQ_DB".CRNT_STEP > 10) AND ("100_BC_AUTO_SEQ_DB".CRNT_STEP < 550)) OR "AlwaysTRUE") AND NOT "10 DI_DATA".FS317 AND NOT "10 DI_DATA".FS320 AND ((NOT "50_CMND_DATA"."TIT 360 Healthy" AND "50_CMND_DATA"."TIT 401 Healthy") OR "50_CMND_DATA"."TIT 360 Healthy");
END_REGION

REGION Network 14: DB62.DBX7.5 = Soot System Power Healthy
   // Word 4 bit 13
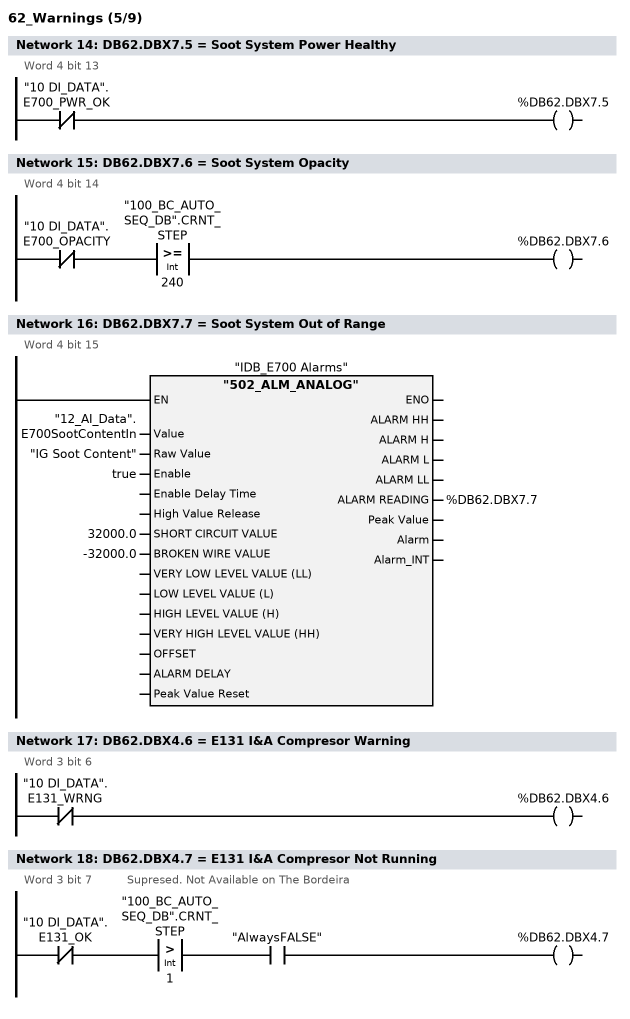
   RUNG wire#powerrail
      I_Contact( "10 DI_DATA".E700_PWR_OK )
      Coil( %DB62.DBX7.5 )
   END_RUNG
   // the same network as SCL:
   %DB62.DBX7.5 := NOT "10 DI_DATA".E700_PWR_OK;
END_REGION
